// folder: State MACHINE/2)Reactors/Reactor R-202/Control R-202

FUNCTION_BLOCK "R-202_Control"   // FB40, GRAPH_PLUS
{ S7_Optimized_Access := 'TRUE' }
VERSION : 0.1
   VAR_INPUT
      OFF_SQ : Bool := false;   // Turn sequence off
      INIT_SQ : Bool := false;   // Set sequence to initial state
      ACK_EF : Bool := false;   // Acknowledge all errors and faults
      "P-201A/B _SEL" : Int := 1;   // IF FALSE P201A is priority / IF TRUE P201B is priority
      "P-202A/B _SEL" : Int := 1;   // IF FALSE P202A is priority / IF TRUE P202B is priority
      IL : Bool;   // INTERLOCKS
   END_VAR
   VAR_OUTPUT
      S_NO : Int := 0;   // Step number
      S_MORE : Bool := false;   // More steps are available and can be shown in S_NO
      S_ACTIVE : Bool := false;   // Step indicated in S_NO is active
      ERR_FLT : Bool := false;   // Interlock or supervision group error
      AUTO_ON : Bool := false;   // Automatic mode is active
   END_VAR
   VAR
      STATE : Int;   // Step number
      Reactor : Struct
         ABORTING : Bool;   // Sequence about
         BatchVolume : Real;   // Batch Volume SP in Liter
         Batchsize : Real;   // Batch size in SP Liter
      END_STRUCT;
      TEMP : Struct
         TANKS_BATCH : Real;   // T-101 & T-102 Batch Sizes
         "EMPTY_LV_0%" : Real;   // 0 % of the Total Batch Size SP
         "MIN_LV_20%" : Real;   // 20 % of the Total Batch Size SP
         "MAX_LV_80%" : Real;   // 80 % of the Total Batch Size SP
         "BELOW_32%" : Real;   // <32% of T-103 Total Batch Size
         "Greater_8%" : Real;   // >8% of T-103 Total Batch Size
         "PRE-ADD" : Real;   // Water & Batch size
         X_SOL_SIZE : Real := 5.0;   // T-101 Soluction Size
         Y_SOL_SIZE : Real := 5.0;   // T-102 Soluction Size
         OFFSEt : Struct
            MAX : Real;
            MIN : Real;
         END_STRUCT;
      END_STRUCT;
      "R-202_TEMP" : Struct
         TANKS_BATCH : Real;   // T-101 & T-102 Batch Sizes
         "EMPTY_LV_0%" : Real;   // 0 % of the Total Batch Size SP
         "MIN_LV_20%" : Real;   // 20 % of the Total Batch Size SP
         "MAX_LV_80%" : Real;   // 80 % of the Total Batch Size SP
         "BELOW_32%" : Real;   // <32% of T-103 Total Batch Size
         "Greater_8%" : Real;   // >8% of T-103 Total Batch Size
         "PRE-ADD" : Real;   // Water & Batch size
         X_SOL_SIZE : Real := 5.0;   // T-101 Soluction Size
         Y_SOL_SIZE : Real := 5.0;   // T-102 Soluction Size
         OFFSEt : Struct
            MAX : Real;
            MIN : Real;
         END_STRUCT;
      END_STRUCT;
      "TIMER" : Array[0..10] of IEC_TIMER;
      "TIME" : Array[0..10] of Time;
      HMI_INFO : Array[0..9] of UInt;
      IF_PAR : G7_IfParPlus_V6;
      RT_DATA : G7_RTDataPlus_V6;   // Internal data area
      Abort : G7_TransitionPlus_V6;   // Transition structure
      "Init R-201" : G7_TransitionPlus_V6;   // Transition structure
      Process : G7_TransitionPlus_V6;   // Transition structure
      TankW : G7_TransitionPlus_V6;   // Transition structure
      TubWash : G7_TransitionPlus_V6;   // Transition structure
      RProcess : G7_TransitionPlus_V6;   // Transition structure
      Trans14 : G7_TransitionPlus_V6;   // Transition structure
      Trans105 : G7_TransitionPlus_V6;   // Transition structure
      Trans106 : G7_TransitionPlus_V6;   // Transition structure
      BachSize : G7_TransitionPlus_V6;   // Transition structure
      Trans110 : G7_TransitionPlus_V6;   // Transition structure
      Trans111 : G7_TransitionPlus_V6;   // Transition structure
      PresetsOK : G7_TransitionPlus_V6;   // Transition structure
      FromHMI : G7_TransitionPlus_V6;   // Transition structure
      Started : G7_TransitionPlus_V6;   // Transition structure
      RDone : G7_TransitionPlus_V6;   // Transition structure
      TDone : G7_TransitionPlus_V6;   // Transition structure
      "R-201 Idle" : G7_TransitionPlus_V6;   // Transition structure
      Trans19 : G7_TransitionPlus_V6;   // Transition structure
      Trans20 : G7_TransitionPlus_V6;   // Transition structure
      TaW : G7_TransitionPlus_V6;   // Transition structure
      TuW : G7_TransitionPlus_V6;   // Transition structure
      DoneAbrt : G7_TransitionPlus_V6;   // Transition structure
      IsIdle : G7_TransitionPlus_V6;   // Transition structure
      Idle : G7_StepPlus_V6;   // Step structure
      Initialize : G7_StepPlus_V6;   // Step structure
      Ready : G7_StepPlus_V6;   // Step structure
      TankWash : G7_StepPlus_V6;   // Step structure
      TubingWash : G7_StepPlus_V6;   // Step structure
      Bach_Size : G7_StepPlus_V6;   // Step structure
      Presets : G7_StepPlus_V6;   // Step structure
      WaitHMI : G7_StepPlus_V6;   // Step structure
      Start : G7_StepPlus_V6;   // Step structure
      Reacting : G7_StepPlus_V6;   // Step structure
      "Transf-->T-103" : G7_StepPlus_V6;   // Step structure
      Done : G7_StepPlus_V6;   // Step structure
      Aborting : G7_StepPlus_V6;   // Step structure
      Release : G7_StepPlus_V6;   // Step structure
      Release_TW : G7_StepPlus_V6;   // Step structure
      Release_TuW : G7_StepPlus_V6;   // Step structure
      RdyTaW : G7_StepPlus_V6;   // Step structure
      RdyTuW : G7_StepPlus_V6;   // Step structure
      SINI : Array[0..2] of USInt;
      LSTT : Array[0..23] of USInt;
      ATAJ : Array[0..23] of USInt;
      ATAB : Array[0..23] of USInt;
      PSTT : Array[0..23] of USInt;
      NSTT : Array[0..23] of USInt;
      ASSJ : Array[0..17] of USInt;
      ASSB : Array[0..17] of USInt;
      PTTS : Array[0..17] of USInt;
      NTTS : Array[0..17] of USInt;
      SW_SQTS : Array[0..17] of USInt;
      SWITCH : Array[0..4] of USInt;
      TVX : Array[0..10] of USInt;
      TTX : Array[0..10] of USInt;
      TSX : Array[0..2] of USInt;
      S00X : Array[0..2] of USInt;
      SOFFX : Array[0..2] of USInt;
      SONX : Array[0..2] of USInt;
      SAX : Array[0..2] of USInt;
      SERRX : Array[0..18] of USInt;
      SMX : Array[0..18] of USInt;
      S0X : Array[0..18] of USInt;
      S1X : Array[0..18] of USInt;
      IL_ALARM_INST : Diag_Alarm;
      SUP_ALARM_INST : Diag_Alarm;
      STEP_TIME_ALARM_INST : Diag_Alarm;
      IEC_TIMER_INST : IEC_TIMER;
      TRANSACTION_FLAG : Bool := false;
   END_VAR
   VAR CONSTANT
      "Single R-201 T-101 seq done" : Int := 214;
      "Single R-201 T-102 seq done" : Int := 218;
   END_VAR
   // SINI[0] := 2;
   // LSTT[0] := 12;
   // NSTT[0] := 12;
   // PTTS[0] := 255;
   // TVX[0] := 16#1;
   // TTX[0] := 16#1;
   // TSX[0] := 16#1;
   // S00X[0] := 16#1;
   // SOFFX[0] := 16#1;
   // SONX[0] := 16#1;
   // SAX[0] := 16#1;
   // SERRX[0] := 16#1;
   // SMX[0] := 16#1;
   // S0X[0] := 16#1;
   // S1X[0] := 16#1;
   // SINI[2] := 255;
   // LSTT[1] := 255;
   // LSTT[2] := 255;
   // LSTT[3] := 255;
   // LSTT[4] := 255;
   // LSTT[5] := 2;
   // LSTT[6] := 255;
   // LSTT[7] := 255;
   // LSTT[8] := 255;
   // LSTT[9] := 255;
   // LSTT[19] := 255;
   // LSTT[12] := 255;
   // LSTT[13] := 255;
   // LSTT[14] := 255;
   // LSTT[15] := 255;
   // LSTT[16] := 255;
   // LSTT[18] := 255;
   // LSTT[20] := 16;
   // LSTT[21] := 17;
   // LSTT[22] := 255;
   // ATAJ[1] := 1;
   // ATAJ[2] := 2;
   // ATAJ[3] := 3;
   // ATAJ[4] := 4;
   // ATAJ[5] := 5;
   // ATAJ[6] := 6;
   // ATAJ[7] := 7;
   // ATAJ[8] := 8;
   // ATAJ[9] := 9;
   // ATAJ[10] := 10;
   // ATAJ[11] := 11;
   // ATAJ[12] := 12;
   // ATAJ[13] := 13;
   // ATAJ[14] := 14;
   // ATAJ[15] := 15;
   // ATAJ[16] := 16;
   // ATAJ[17] := 17;
   // ATAJ[18] := 18;
   // ATAJ[19] := 19;
   // ATAJ[20] := 20;
   // ATAJ[21] := 21;
   // ATAJ[22] := 22;
   // ATAJ[23] := 23;
   // ATAB[1] := 2;
   // ATAB[2] := 3;
   // ATAB[3] := 4;
   // ATAB[20] := 21;
   // ATAB[5] := 20;
   // ATAB[6] := 6;
   // ATAB[7] := 7;
   // ATAB[8] := 8;
   // ATAB[9] := 9;
   // ATAB[10] := 10;
   // ATAB[11] := 11;
   // ATAB[12] := 12;
   // ATAB[13] := 13;
   // ATAB[14] := 14;
   // ATAB[15] := 15;
   // ATAB[16] := 16;
   // ATAB[17] := 17;
   // ATAB[18] := 18;
   // ATAB[19] := 19;
   // ATAB[21] := 5;
   // ATAB[22] := 22;
   // ATAB[23] := 23;
   // PSTT[20] := 1;
   // PSTT[5] := 1;
   // PSTT[6] := 2;
   // PSTT[7] := 3;
   // PSTT[8] := 4;
   // PSTT[9] := 5;
   // PSTT[10] := 14;
   // PSTT[11] := 15;
   // PSTT[12] := 6;
   // PSTT[13] := 7;
   // PSTT[14] := 8;
   // PSTT[15] := 9;
   // PSTT[16] := 10;
   // PSTT[17] := 11;
   // PSTT[18] := 16;
   // PSTT[19] := 17;
   // PSTT[21] := 1;
   // PSTT[22] := 12;
   // PSTT[23] := 13;
   // NSTT[1] := 1;
   // NSTT[2] := 2;
   // NSTT[3] := 16;
   // NSTT[4] := 17;
   // NSTT[5] := 2;
   // NSTT[6] := 5;
   // NSTT[7] := 14;
   // NSTT[8] := 15;
   // NSTT[9] := 6;
   // NSTT[19] := 4;
   // NSTT[12] := 7;
   // NSTT[13] := 8;
   // NSTT[14] := 9;
   // NSTT[15] := 10;
   // NSTT[16] := 11;
   // NSTT[18] := 3;
   // NSTT[20] := 16;
   // NSTT[21] := 17;
   // NSTT[22] := 13;
   // ASSJ[1] := 1;
   // ASSJ[2] := 2;
   // ASSJ[3] := 3;
   // ASSJ[4] := 4;
   // ASSJ[5] := 5;
   // ASSJ[6] := 6;
   // ASSJ[7] := 7;
   // ASSJ[8] := 8;
   // ASSJ[9] := 9;
   // ASSJ[10] := 10;
   // ASSJ[11] := 11;
   // ASSJ[12] := 12;
   // ASSJ[13] := 13;
   // ASSJ[14] := 14;
   // ASSJ[15] := 15;
   // ASSJ[16] := 16;
   // ASSJ[17] := 17;
   // ASSB[1] := 1;
   // ASSB[2] := 2;
   // ASSB[3] := 3;
   // ASSB[4] := 4;
   // ASSB[5] := 5;
   // ASSB[6] := 6;
   // ASSB[7] := 7;
   // ASSB[8] := 8;
   // ASSB[9] := 9;
   // ASSB[10] := 10;
   // ASSB[11] := 11;
   // ASSB[12] := 12;
   // ASSB[13] := 13;
   // ASSB[14] := 14;
   // ASSB[15] := 15;
   // ASSB[16] := 16;
   // ASSB[17] := 17;
   // PTTS[2] := 2;
   // PTTS[3] := 18;
   // PTTS[4] := 19;
   // PTTS[5] := 6;
   // PTTS[6] := 9;
   // PTTS[7] := 12;
   // PTTS[8] := 13;
   // PTTS[9] := 14;
   // PTTS[10] := 15;
   // PTTS[11] := 16;
   // PTTS[12] := 255;
   // PTTS[13] := 22;
   // PTTS[14] := 7;
   // PTTS[16] := 3;
   // PTTS[17] := 4;
   // PTTS[15] := 8;
   // NTTS[1] := 5;
   // NTTS[2] := 6;
   // NTTS[3] := 7;
   // NTTS[4] := 8;
   // NTTS[5] := 9;
   // NTTS[6] := 12;
   // NTTS[7] := 13;
   // NTTS[8] := 14;
   // NTTS[9] := 15;
   // NTTS[10] := 16;
   // NTTS[11] := 17;
   // NTTS[12] := 22;
   // NTTS[13] := 23;
   // NTTS[14] := 10;
   // NTTS[15] := 11;
   // NTTS[16] := 18;
   // NTTS[17] := 19;
   // SW_SQTS[2] := 2;
   // SW_SQTS[3] := 3;
   // SW_SQTS[4] := 4;
   // SW_SQTS[5] := 2;
   // SW_SQTS[6] := 2;
   // SW_SQTS[7] := 2;
   // SW_SQTS[8] := 2;
   // SW_SQTS[9] := 2;
   // SW_SQTS[10] := 2;
   // SW_SQTS[11] := 2;
   // SW_SQTS[12] := 5;
   // SW_SQTS[13] := 5;
   // SW_SQTS[14] := 3;
   // SW_SQTS[15] := 4;
   // SW_SQTS[16] := 3;
   // SW_SQTS[17] := 4;
   // SWITCH[1] := 8;
   // SWITCH[2] := 130;
   // SWITCH[3] := 224;
   // SWITCH[4] := 7;
   // ATAB[0] := 1;
   // PTTS[1] := 1;
   // SW_SQTS[1] := 1;
   // SWITCH[0] := 32;
BEGIN
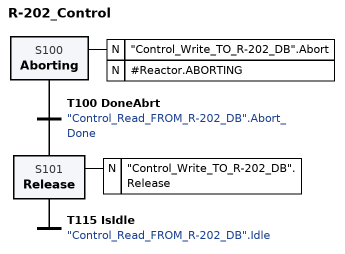
   // sequencer 1
   STEP Aborting:   // S100, max time T#10S, warning time T#7S
      // T-101 Pouring Soluction Valve
              N    "Control_Write_TO_R-202_DB".Abort
              N    #Reactor.ABORTING
   END_STEP
   TRANSITION DoneAbrt FROM Aborting TO Release   // T100: CLOSED: XV-1041 XV-1011 XV-1013OFF: VFD-1011 P-101A P-101BZERO: FT-1041 Totalizer
      := "Control_Read_FROM_R-202_DB".Abort_Done;
   END_TRANSITION
   STEP Release:   // S101, max time T#10S, warning time T#7S
              N    "Control_Write_TO_R-202_DB".Release
   END_STEP
   TRANSITION IsIdle FROM Release TO ?   // T115
      := "Control_Read_FROM_R-202_DB".Idle;
   END_TRANSITION
END_FUNCTION_BLOCK

FUNCTION "R-202_CTRL_SEQ_FC" : Void   // FC44, LAD
{ S7_Optimized_Access := 'TRUE' }
VERSION : 0.1
   VAR_TEMP   // added for the SCL form of the ladder/FBD networks
      _w1 : Bool;
   END_VAR
BEGIN

REGION Network 2: Reset Abort Cmd
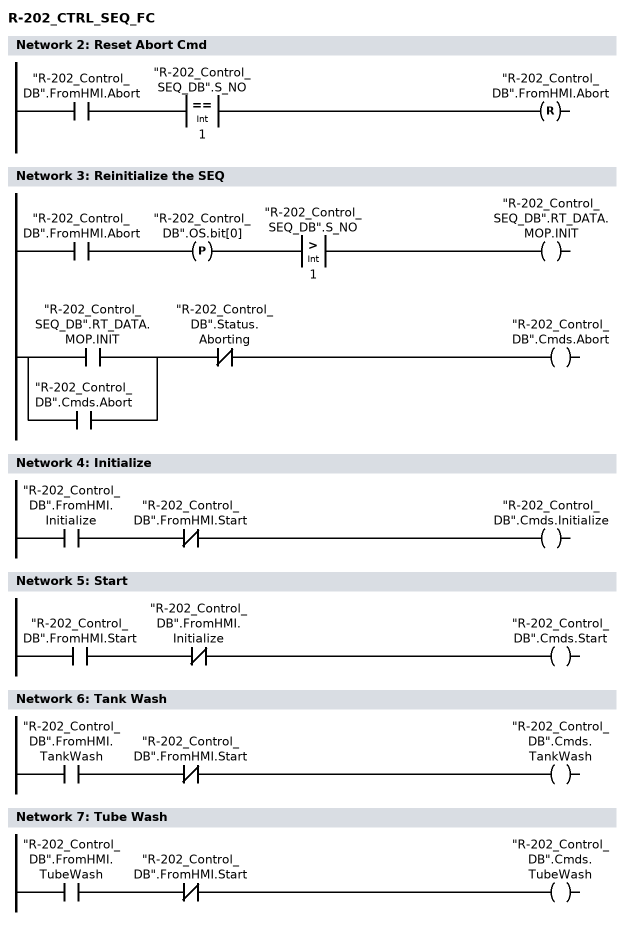
   RUNG wire#powerrail
      Contact( "R-202_Control_DB".FromHMI.Abort )
      { S7_Templates := "SrcType := Int" } EQ_Contact(in1 := "R-202_Control_SEQ_DB".S_NO, in2 := 1)
      R_Coil( "R-202_Control_DB".FromHMI.Abort )
   END_RUNG
   // the same network as SCL:
   IF "R-202_Control_DB".FromHMI.Abort AND ("R-202_Control_SEQ_DB".S_NO = 1) THEN
       "R-202_Control_DB".FromHMI.Abort := FALSE;
   END_IF;
END_REGION

REGION Network 3: Reinitialize the SEQ
   RUNG wire#powerrail
      Contact( "R-202_Control_DB".FromHMI.Abort )
      P_Trig( "R-202_Control_DB".OS.bit[0] )
      { S7_Templates := "SrcType := Int" } GT_Contact(in1 := "R-202_Control_SEQ_DB".S_NO, in2 := 1)
      Coil( "R-202_Control_SEQ_DB".RT_DATA.MOP.INIT )
   END_RUNG
   RUNG wire#powerrail
      Contact( "R-202_Control_SEQ_DB".RT_DATA.MOP.INIT )
      wire#w1
      I_Contact( "R-202_Control_DB".Status.Aborting )
      Coil( "R-202_Control_DB".Cmds.Abort )
   END_RUNG
   RUNG wire#powerrail
      Contact( "R-202_Control_DB".Cmds.Abort )
   END_RUNG wire#w1
   // the same network as SCL:
   #_w1 := "R-202_Control_DB".FromHMI.Abort AND NOT "R-202_Control_DB".OS.bit[0];   // rising edge
   "R-202_Control_DB".OS.bit[0] := "R-202_Control_DB".FromHMI.Abort;
   "R-202_Control_SEQ_DB".RT_DATA.MOP.INIT := #_w1 AND ("R-202_Control_SEQ_DB".S_NO > 1);
   "R-202_Control_DB".Cmds.Abort := ("R-202_Control_SEQ_DB".RT_DATA.MOP.INIT OR "R-202_Control_DB".Cmds.Abort) AND NOT "R-202_Control_DB".Status.Aborting;
END_REGION

REGION Network 4: Initialize
   RUNG wire#powerrail
      Contact( "R-202_Control_DB".FromHMI.Initialize )
      I_Contact( "R-202_Control_DB".FromHMI.Start )
      Coil( "R-202_Control_DB".Cmds.Initialize )
   END_RUNG
   // the same network as SCL:
   "R-202_Control_DB".Cmds.Initialize := "R-202_Control_DB".FromHMI.Initialize AND NOT "R-202_Control_DB".FromHMI.Start;
END_REGION

REGION Network 5: Start
   RUNG wire#powerrail
      Contact( "R-202_Control_DB".FromHMI.Start )
      I_Contact( "R-202_Control_DB".FromHMI.Initialize )
      Coil( "R-202_Control_DB".Cmds.Start )
   END_RUNG
   // the same network as SCL:
   "R-202_Control_DB".Cmds.Start := "R-202_Control_DB".FromHMI.Start AND NOT "R-202_Control_DB".FromHMI.Initialize;
END_REGION

REGION Network 6: Tank Wash
   RUNG wire#powerrail
      Contact( "R-202_Control_DB".FromHMI.TankWash )
      I_Contact( "R-202_Control_DB".FromHMI.Start )
      Coil( "R-202_Control_DB".Cmds.TankWash )
   END_RUNG
   // the same network as SCL:
   "R-202_Control_DB".Cmds.TankWash := "R-202_Control_DB".FromHMI.TankWash AND NOT "R-202_Control_DB".FromHMI.Start;
END_REGION

REGION Network 7: Tube Wash
   RUNG wire#powerrail
      Contact( "R-202_Control_DB".FromHMI.TubeWash )
      I_Contact( "R-202_Control_DB".FromHMI.Start )
      Coil( "R-202_Control_DB".Cmds.TubeWash )
   END_RUNG
   // the same network as SCL:
   "R-202_Control_DB".Cmds.TubeWash := "R-202_Control_DB".FromHMI.TubeWash AND NOT "R-202_Control_DB".FromHMI.Start;
END_REGION
END_FUNCTION

// folder: State MACHINE/2)Reactors/Reactor R-202/Control R-202/Control <---> R-202

FUNCTION "Control_Signals_FROM_R-202" : Void   // FC54, LAD
{ S7_Optimized_Access := 'TRUE' }
VERSION : 0.1
BEGIN

REGION Network 1: R-201 Initialization Done
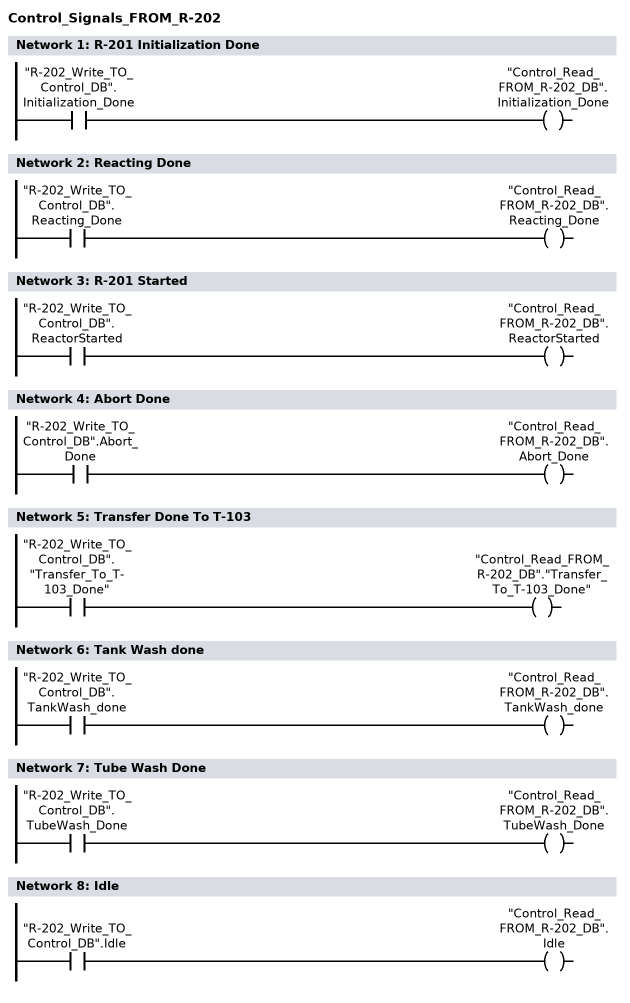
   RUNG wire#powerrail
      Contact( "R-202_Write_TO_Control_DB".Initialization_Done )
      Coil( "Control_Read_FROM_R-202_DB".Initialization_Done )
   END_RUNG
   // the same network as SCL:
   "Control_Read_FROM_R-202_DB".Initialization_Done := "R-202_Write_TO_Control_DB".Initialization_Done;
END_REGION

REGION Network 2: Reacting Done
   RUNG wire#powerrail
      Contact( "R-202_Write_TO_Control_DB".Reacting_Done )
      Coil( "Control_Read_FROM_R-202_DB".Reacting_Done )
   END_RUNG
   // the same network as SCL:
   "Control_Read_FROM_R-202_DB".Reacting_Done := "R-202_Write_TO_Control_DB".Reacting_Done;
END_REGION

REGION Network 3: R-201 Started
   RUNG wire#powerrail
      Contact( "R-202_Write_TO_Control_DB".ReactorStarted )
      Coil( "Control_Read_FROM_R-202_DB".ReactorStarted )
   END_RUNG
   // the same network as SCL:
   "Control_Read_FROM_R-202_DB".ReactorStarted := "R-202_Write_TO_Control_DB".ReactorStarted;
END_REGION

REGION Network 4: Abort Done
   RUNG wire#powerrail
      Contact( "R-202_Write_TO_Control_DB".Abort_Done )
      Coil( "Control_Read_FROM_R-202_DB".Abort_Done )
   END_RUNG
   // the same network as SCL:
   "Control_Read_FROM_R-202_DB".Abort_Done := "R-202_Write_TO_Control_DB".Abort_Done;
END_REGION

REGION Network 5: Transfer Done To T-103
   RUNG wire#powerrail
      Contact( "R-202_Write_TO_Control_DB"."Transfer_To_T-103_Done" )
      Coil( "Control_Read_FROM_R-202_DB"."Transfer_To_T-103_Done" )
   END_RUNG
   // the same network as SCL:
   "Control_Read_FROM_R-202_DB"."Transfer_To_T-103_Done" := "R-202_Write_TO_Control_DB"."Transfer_To_T-103_Done";
END_REGION

REGION Network 6: Tank Wash done
   RUNG wire#powerrail
      Contact( "R-202_Write_TO_Control_DB".TankWash_done )
      Coil( "Control_Read_FROM_R-202_DB".TankWash_done )
   END_RUNG
   // the same network as SCL:
   "Control_Read_FROM_R-202_DB".TankWash_done := "R-202_Write_TO_Control_DB".TankWash_done;
END_REGION

REGION Network 7: Tube Wash Done
   RUNG wire#powerrail
      Contact( "R-202_Write_TO_Control_DB".TubeWash_Done )
      Coil( "Control_Read_FROM_R-202_DB".TubeWash_Done )
   END_RUNG
   // the same network as SCL:
   "Control_Read_FROM_R-202_DB".TubeWash_Done := "R-202_Write_TO_Control_DB".TubeWash_Done;
END_REGION

REGION Network 8: Idle
   RUNG wire#powerrail
      Contact( "R-202_Write_TO_Control_DB".Idle )
      Coil( "Control_Read_FROM_R-202_DB".Idle )
   END_RUNG
   // the same network as SCL:
   "Control_Read_FROM_R-202_DB".Idle := "R-202_Write_TO_Control_DB".Idle;
END_REGION
END_FUNCTION

// folder: State MACHINE/2)Reactors/Reactor R-202/R-202 <---> Control

FUNCTION "R-202_Signals_FROM_Control" : Void   // FC47, LAD
{ S7_Optimized_Access := 'TRUE' }
VERSION : 0.1
BEGIN

REGION Network 1: Start From Reactor Selector.
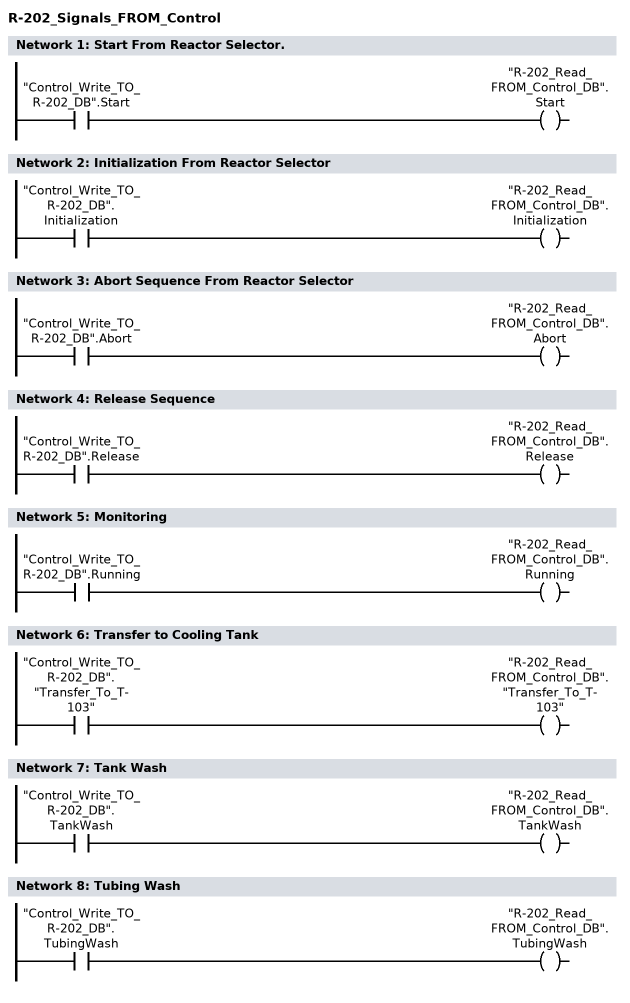
   RUNG wire#powerrail
      Contact( "Control_Write_TO_R-202_DB".Start )
      Coil( "R-202_Read_FROM_Control_DB".Start )
   END_RUNG
   // the same network as SCL:
   "R-202_Read_FROM_Control_DB".Start := "Control_Write_TO_R-202_DB".Start;
END_REGION

REGION Network 2: Initialization From Reactor Selector
   RUNG wire#powerrail
      Contact( "Control_Write_TO_R-202_DB".Initialization )
      Coil( "R-202_Read_FROM_Control_DB".Initialization )
   END_RUNG
   // the same network as SCL:
   "R-202_Read_FROM_Control_DB".Initialization := "Control_Write_TO_R-202_DB".Initialization;
END_REGION

REGION Network 3: Abort Sequence From Reactor Selector
   RUNG wire#powerrail
      Contact( "Control_Write_TO_R-202_DB".Abort )
      Coil( "R-202_Read_FROM_Control_DB".Abort )
   END_RUNG
   // the same network as SCL:
   "R-202_Read_FROM_Control_DB".Abort := "Control_Write_TO_R-202_DB".Abort;
END_REGION

REGION Network 4: Release Sequence
   RUNG wire#powerrail
      Contact( "Control_Write_TO_R-202_DB".Release )
      Coil( "R-202_Read_FROM_Control_DB".Release )
   END_RUNG
   // the same network as SCL:
   "R-202_Read_FROM_Control_DB".Release := "Control_Write_TO_R-202_DB".Release;
END_REGION

REGION Network 5: Monitoring
   RUNG wire#powerrail
      Contact( "Control_Write_TO_R-202_DB".Running )
      Coil( "R-202_Read_FROM_Control_DB".Running )
   END_RUNG
   // the same network as SCL:
   "R-202_Read_FROM_Control_DB".Running := "Control_Write_TO_R-202_DB".Running;
END_REGION

REGION Network 6: Transfer to Cooling Tank
   RUNG wire#powerrail
      Contact( "Control_Write_TO_R-202_DB"."Transfer_To_T-103" )
      Coil( "R-202_Read_FROM_Control_DB"."Transfer_To_T-103" )
   END_RUNG
   // the same network as SCL:
   "R-202_Read_FROM_Control_DB"."Transfer_To_T-103" := "Control_Write_TO_R-202_DB"."Transfer_To_T-103";
END_REGION

REGION Network 7: Tank Wash
   RUNG wire#powerrail
      Contact( "Control_Write_TO_R-202_DB".TankWash )
      Coil( "R-202_Read_FROM_Control_DB".TankWash )
   END_RUNG
   // the same network as SCL:
   "R-202_Read_FROM_Control_DB".TankWash := "Control_Write_TO_R-202_DB".TankWash;
END_REGION

REGION Network 8: Tubing Wash
   RUNG wire#powerrail
      Contact( "Control_Write_TO_R-202_DB".TubingWash )
      Coil( "R-202_Read_FROM_Control_DB".TubingWash )
   END_RUNG
   // the same network as SCL:
   "R-202_Read_FROM_Control_DB".TubingWash := "Control_Write_TO_R-202_DB".TubingWash;
END_REGION
END_FUNCTION

// folder: State MACHINE/2)Reactors/Reactor R-202/R-202 <---> T-101

FUNCTION "R-202_Signals_FROM_T-101" : Void   // FC62, LAD
{ S7_Optimized_Access := 'TRUE' }
VERSION : 0.1
BEGIN

REGION Network 1: Start Sequence
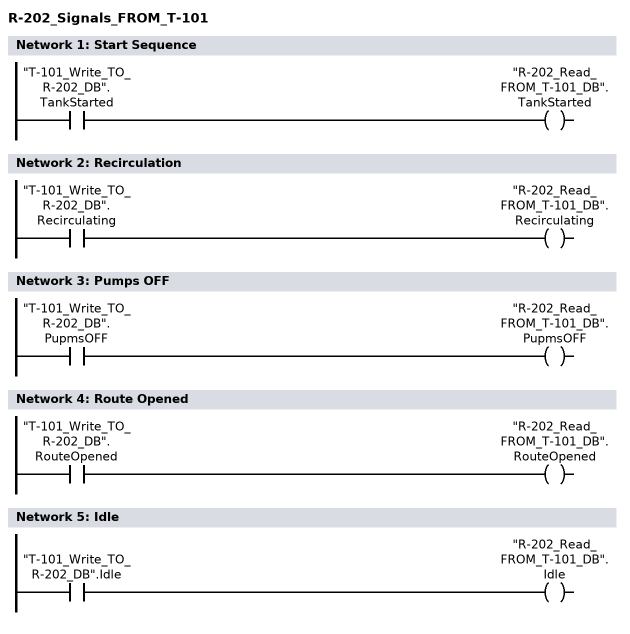
   RUNG wire#powerrail
      Contact( "T-101_Write_TO_R-202_DB".TankStarted )
      Coil( "R-202_Read_FROM_T-101_DB".TankStarted )
   END_RUNG
   // the same network as SCL:
   "R-202_Read_FROM_T-101_DB".TankStarted := "T-101_Write_TO_R-202_DB".TankStarted;
END_REGION

REGION Network 2: Recirculation
   RUNG wire#powerrail
      Contact( "T-101_Write_TO_R-202_DB".Recirculating )
      Coil( "R-202_Read_FROM_T-101_DB".Recirculating )
   END_RUNG
   // the same network as SCL:
   "R-202_Read_FROM_T-101_DB".Recirculating := "T-101_Write_TO_R-202_DB".Recirculating;
END_REGION

REGION Network 3: Pumps OFF
   RUNG wire#powerrail
      Contact( "T-101_Write_TO_R-202_DB".PupmsOFF )
      Coil( "R-202_Read_FROM_T-101_DB".PupmsOFF )
   END_RUNG
   // the same network as SCL:
   "R-202_Read_FROM_T-101_DB".PupmsOFF := "T-101_Write_TO_R-202_DB".PupmsOFF;
END_REGION

REGION Network 4: Route Opened
   RUNG wire#powerrail
      Contact( "T-101_Write_TO_R-202_DB".RouteOpened )
      Coil( "R-202_Read_FROM_T-101_DB".RouteOpened )
   END_RUNG
   // the same network as SCL:
   "R-202_Read_FROM_T-101_DB".RouteOpened := "T-101_Write_TO_R-202_DB".RouteOpened;
END_REGION

REGION Network 5: Idle
   RUNG wire#powerrail
      Contact( "T-101_Write_TO_R-202_DB".Idle )
      Coil( "R-202_Read_FROM_T-101_DB".Idle )
   END_RUNG
   // the same network as SCL:
   "R-202_Read_FROM_T-101_DB".Idle := "T-101_Write_TO_R-202_DB".Idle;
END_REGION
END_FUNCTION

// folder: State MACHINE/2)Reactors/Reactor R-202/R-202 <---> T-102

FUNCTION "R-202_Signals_FROM_T-102" : Void   // FC59, LAD
{ S7_Optimized_Access := 'TRUE' }
VERSION : 0.1
BEGIN

REGION Network 1: Start Sequence
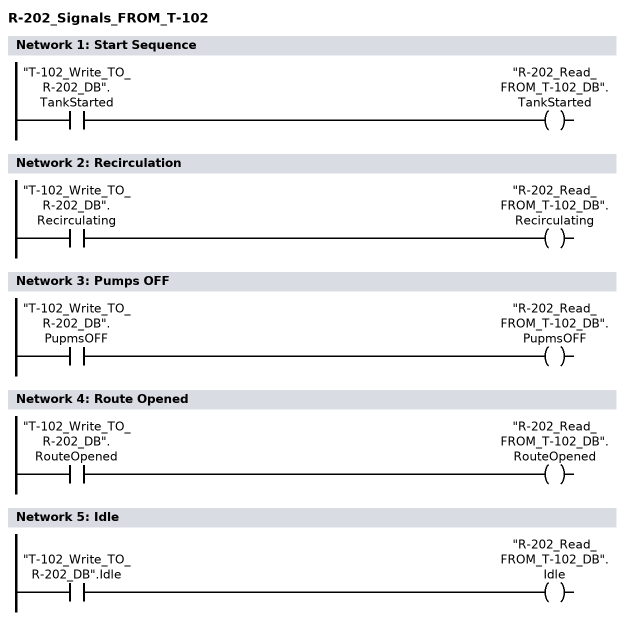
   RUNG wire#powerrail
      Contact( "T-102_Write_TO_R-202_DB".TankStarted )
      Coil( "R-202_Read_FROM_T-102_DB".TankStarted )
   END_RUNG
   // the same network as SCL:
   "R-202_Read_FROM_T-102_DB".TankStarted := "T-102_Write_TO_R-202_DB".TankStarted;
END_REGION

REGION Network 2: Recirculation
   RUNG wire#powerrail
      Contact( "T-102_Write_TO_R-202_DB".Recirculating )
      Coil( "R-202_Read_FROM_T-102_DB".Recirculating )
   END_RUNG
   // the same network as SCL:
   "R-202_Read_FROM_T-102_DB".Recirculating := "T-102_Write_TO_R-202_DB".Recirculating;
END_REGION

REGION Network 3: Pumps OFF
   RUNG wire#powerrail
      Contact( "T-102_Write_TO_R-202_DB".PupmsOFF )
      Coil( "R-202_Read_FROM_T-102_DB".PupmsOFF )
   END_RUNG
   // the same network as SCL:
   "R-202_Read_FROM_T-102_DB".PupmsOFF := "T-102_Write_TO_R-202_DB".PupmsOFF;
END_REGION

REGION Network 4: Route Opened
   RUNG wire#powerrail
      Contact( "T-102_Write_TO_R-202_DB".RouteOpened )
      Coil( "R-202_Read_FROM_T-102_DB".RouteOpened )
   END_RUNG
   // the same network as SCL:
   "R-202_Read_FROM_T-102_DB".RouteOpened := "T-102_Write_TO_R-202_DB".RouteOpened;
END_REGION

REGION Network 5: Idle
   RUNG wire#powerrail
      Contact( "T-102_Write_TO_R-202_DB".Idle )
      Coil( "R-202_Read_FROM_T-102_DB".Idle )
   END_RUNG
   // the same network as SCL:
   "R-202_Read_FROM_T-102_DB".Idle := "T-102_Write_TO_R-202_DB".Idle;
END_REGION
END_FUNCTION

// folder: State MACHINE/2)Reactors/Reactor R-202/R-202 <---> T-103 (CoolingTank)

FUNCTION "R-202_Signals_FROM_T-103" : Void   // FC58, LAD
{ S7_Optimized_Access := 'TRUE' }
VERSION : 0.1
BEGIN

REGION Network 1: Start Sequence
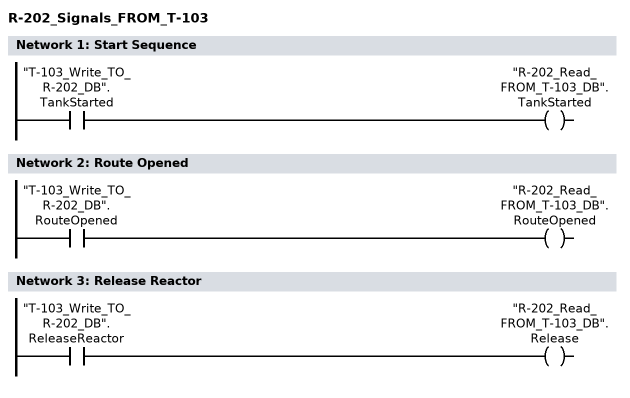
   RUNG wire#powerrail
      Contact( "T-103_Write_TO_R-202_DB".TankStarted )
      Coil( "R-202_Read_FROM_T-103_DB".TankStarted )
   END_RUNG
   // the same network as SCL:
   "R-202_Read_FROM_T-103_DB".TankStarted := "T-103_Write_TO_R-202_DB".TankStarted;
END_REGION

REGION Network 2: Route Opened
   RUNG wire#powerrail
      Contact( "T-103_Write_TO_R-202_DB".RouteOpened )
      Coil( "R-202_Read_FROM_T-103_DB".RouteOpened )
   END_RUNG
   // the same network as SCL:
   "R-202_Read_FROM_T-103_DB".RouteOpened := "T-103_Write_TO_R-202_DB".RouteOpened;
END_REGION

REGION Network 3: Release Reactor
   RUNG wire#powerrail
      Contact( "T-103_Write_TO_R-202_DB".ReleaseReactor )
      Coil( "R-202_Read_FROM_T-103_DB".Release )
   END_RUNG
   // the same network as SCL:
   "R-202_Read_FROM_T-103_DB".Release := "T-103_Write_TO_R-202_DB".ReleaseReactor;
END_REGION
END_FUNCTION

// folder: State MACHINE/2)Reactors/Reactor R-202/R-202 <---> T-104 (WaterSystem)

FUNCTION "R-202_Signals_FROM_T-104" : Void   // FC57, LAD
{ S7_Optimized_Access := 'TRUE' }
VERSION : 0.1
BEGIN

REGION Network 1: Start Sequence
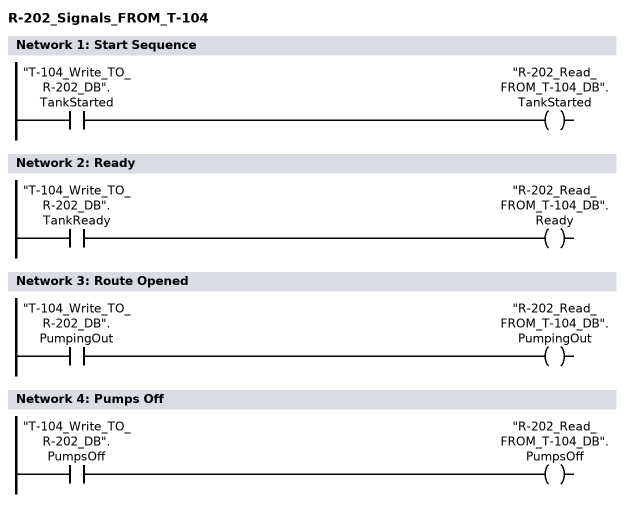
   RUNG wire#powerrail
      Contact( "T-104_Write_TO_R-202_DB".TankStarted )
      Coil( "R-202_Read_FROM_T-104_DB".TankStarted )
   END_RUNG
   // the same network as SCL:
   "R-202_Read_FROM_T-104_DB".TankStarted := "T-104_Write_TO_R-202_DB".TankStarted;
END_REGION

REGION Network 2: Ready
   RUNG wire#powerrail
      Contact( "T-104_Write_TO_R-202_DB".TankReady )
      Coil( "R-202_Read_FROM_T-104_DB".Ready )
   END_RUNG
   // the same network as SCL:
   "R-202_Read_FROM_T-104_DB".Ready := "T-104_Write_TO_R-202_DB".TankReady;
END_REGION

REGION Network 3: Route Opened
   RUNG wire#powerrail
      Contact( "T-104_Write_TO_R-202_DB".PumpingOut )
      Coil( "R-202_Read_FROM_T-104_DB".PumpingOut )
   END_RUNG
   // the same network as SCL:
   "R-202_Read_FROM_T-104_DB".PumpingOut := "T-104_Write_TO_R-202_DB".PumpingOut;
END_REGION

REGION Network 4: Pumps Off
   RUNG wire#powerrail
      Contact( "T-104_Write_TO_R-202_DB".PumpsOff )
      Coil( "R-202_Read_FROM_T-104_DB".PumpsOff )
   END_RUNG
   // the same network as SCL:
   "R-202_Read_FROM_T-104_DB".PumpsOff := "T-104_Write_TO_R-202_DB".PumpsOff;
END_REGION
END_FUNCTION

// folder: State MACHINE/3)Centrifuge

FUNCTION_BLOCK "Centrifuge_SEQ"   // FB28, GRAPH_PLUS
{ S7_Optimized_Access := 'TRUE' }